REGION Network 339: CARRIER SPACING FAULT
   RUNG wire#powerrail
      Contact( "reset" )
      Contact( "EMS".Carrier[59].SDC_OUT.Faults.CarrierSpacingFault )
      wire#w1
      Coil( "DB302_HMI_Faults".Carrier59_Faults_2.%X2 )
   END_RUNG
   RUNG wire#powerrail
      Contact( "DB302_HMI_Faults".Carrier59_Faults_2.%X2 )
      I_Contact( "EMS_Fault_Reset" )
   END_RUNG wire#w1
   // the same network as SCL:
   "DB302_HMI_Faults".Carrier59_Faults_2.%X2 := ("reset" AND "EMS".Carrier[59].SDC_OUT.Faults.CarrierSpacingFault) OR ("DB302_HMI_Faults".Carrier59_Faults_2.%X2 AND NOT "EMS_Fault_Reset");
END_REGION

REGION Network 340: DUPLICATE CARRIER NUMBER FAULT
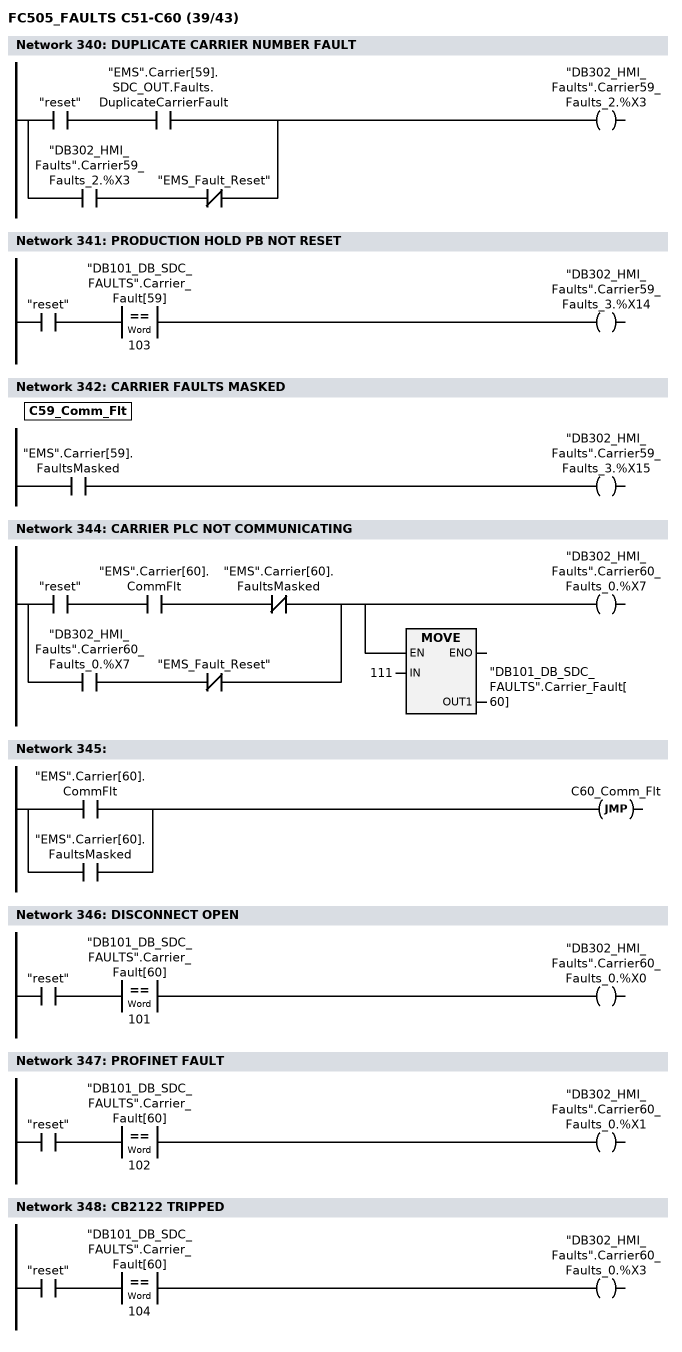
   RUNG wire#powerrail
      Contact( "reset" )
      Contact( "EMS".Carrier[59].SDC_OUT.Faults.DuplicateCarrierFault )
      wire#w1
      Coil( "DB302_HMI_Faults".Carrier59_Faults_2.%X3 )
   END_RUNG
   RUNG wire#powerrail
      Contact( "DB302_HMI_Faults".Carrier59_Faults_2.%X3 )
      I_Contact( "EMS_Fault_Reset" )
   END_RUNG wire#w1
   // the same network as SCL:
   "DB302_HMI_Faults".Carrier59_Faults_2.%X3 := ("reset" AND "EMS".Carrier[59].SDC_OUT.Faults.DuplicateCarrierFault) OR ("DB302_HMI_Faults".Carrier59_Faults_2.%X3 AND NOT "EMS_Fault_Reset");
END_REGION

REGION Network 341: PRODUCTION HOLD PB NOT RESET
   RUNG wire#powerrail
      Contact( "reset" )
      { S7_Templates := "SrcType := Word" } EQ_Contact(in1 := "DB101_DB_SDC_FAULTS".Carrier_Fault[59], in2 := 103)
      Coil( "DB302_HMI_Faults".Carrier59_Faults_3.%X14 )
   END_RUNG
   // the same network as SCL:
   "DB302_HMI_Faults".Carrier59_Faults_3.%X14 := "reset" AND ("DB101_DB_SDC_FAULTS".Carrier_Fault[59] = 103);
END_REGION

REGION Network 342: CARRIER FAULTS MASKED
   Label( C59_Comm_Flt )
   RUNG wire#powerrail
      Contact( "EMS".Carrier[59].FaultsMasked )
      Coil( "DB302_HMI_Faults".Carrier59_Faults_3.%X15 )
   END_RUNG
   // the same network as SCL:
   C59_Comm_Flt:
   "DB302_HMI_Faults".Carrier59_Faults_3.%X15 := "EMS".Carrier[59].FaultsMasked;
END_REGION

REGION Network 343: CARRIER 60 FAULTS
END_REGION

REGION Network 344: CARRIER PLC NOT COMMUNICATING
   RUNG wire#powerrail
      Contact( "reset" )
      Contact( "EMS".Carrier[60].CommFlt )
      I_Contact( "EMS".Carrier[60].FaultsMasked )
      wire#w1
      Coil( "DB302_HMI_Faults".Carrier60_Faults_0.%X7 )
   END_RUNG
   RUNG wire#powerrail
      Contact( "DB302_HMI_Faults".Carrier60_Faults_0.%X7 )
      I_Contact( "EMS_Fault_Reset" )
   END_RUNG wire#w1
   RUNG wire#w1
      Move(in := 111, out1 => "DB101_DB_SDC_FAULTS".Carrier_Fault[60])
   END_RUNG
   // the same network as SCL:
   "DB302_HMI_Faults".Carrier60_Faults_0.%X7 := ("reset" AND "EMS".Carrier[60].CommFlt AND NOT "EMS".Carrier[60].FaultsMasked) OR ("DB302_HMI_Faults".Carrier60_Faults_0.%X7 AND NOT "EMS_Fault_Reset");
   IF "DB302_HMI_Faults".Carrier60_Faults_0.%X7 THEN "DB101_DB_SDC_FAULTS".Carrier_Fault[60] := 111; END_IF;
END_REGION

REGION Network 345
   RUNG wire#powerrail
      Contact( "EMS".Carrier[60].CommFlt )
      wire#w1
      JumpCoil( C60_Comm_Flt )
   END_RUNG
   RUNG wire#powerrail
      Contact( "EMS".Carrier[60].FaultsMasked )
   END_RUNG wire#w1
   // the same network as SCL:
   IF "EMS".Carrier[60].CommFlt OR "EMS".Carrier[60].FaultsMasked THEN GOTO C60_Comm_Flt; END_IF;
END_REGION

REGION Network 346: DISCONNECT OPEN
   RUNG wire#powerrail
      Contact( "reset" )
      { S7_Templates := "SrcType := Word" } EQ_Contact(in1 := "DB101_DB_SDC_FAULTS".Carrier_Fault[60], in2 := 101)
      Coil( "DB302_HMI_Faults".Carrier60_Faults_0.%X0 )
   END_RUNG
   // the same network as SCL:
   "DB302_HMI_Faults".Carrier60_Faults_0.%X0 := "reset" AND ("DB101_DB_SDC_FAULTS".Carrier_Fault[60] = 101);
END_REGION

REGION Network 347: PROFINET FAULT
   RUNG wire#powerrail
      Contact( "reset" )
      { S7_Templates := "SrcType := Word" } EQ_Contact(in1 := "DB101_DB_SDC_FAULTS".Carrier_Fault[60], in2 := 102)
      Coil( "DB302_HMI_Faults".Carrier60_Faults_0.%X1 )
   END_RUNG
   // the same network as SCL:
   "DB302_HMI_Faults".Carrier60_Faults_0.%X1 := "reset" AND ("DB101_DB_SDC_FAULTS".Carrier_Fault[60] = 102);
END_REGION

REGION Network 348: CB2122 TRIPPED
   RUNG wire#powerrail
      Contact( "reset" )
      { S7_Templates := "SrcType := Word" } EQ_Contact(in1 := "DB101_DB_SDC_FAULTS".Carrier_Fault[60], in2 := 104)
      Coil( "DB302_HMI_Faults".Carrier60_Faults_0.%X3 )
   END_RUNG
   // the same network as SCL:
   "DB302_HMI_Faults".Carrier60_Faults_0.%X3 := "reset" AND ("DB101_DB_SDC_FAULTS".Carrier_Fault[60] = 104);
END_REGION

REGION Network 349: CB2123 TRIPPED
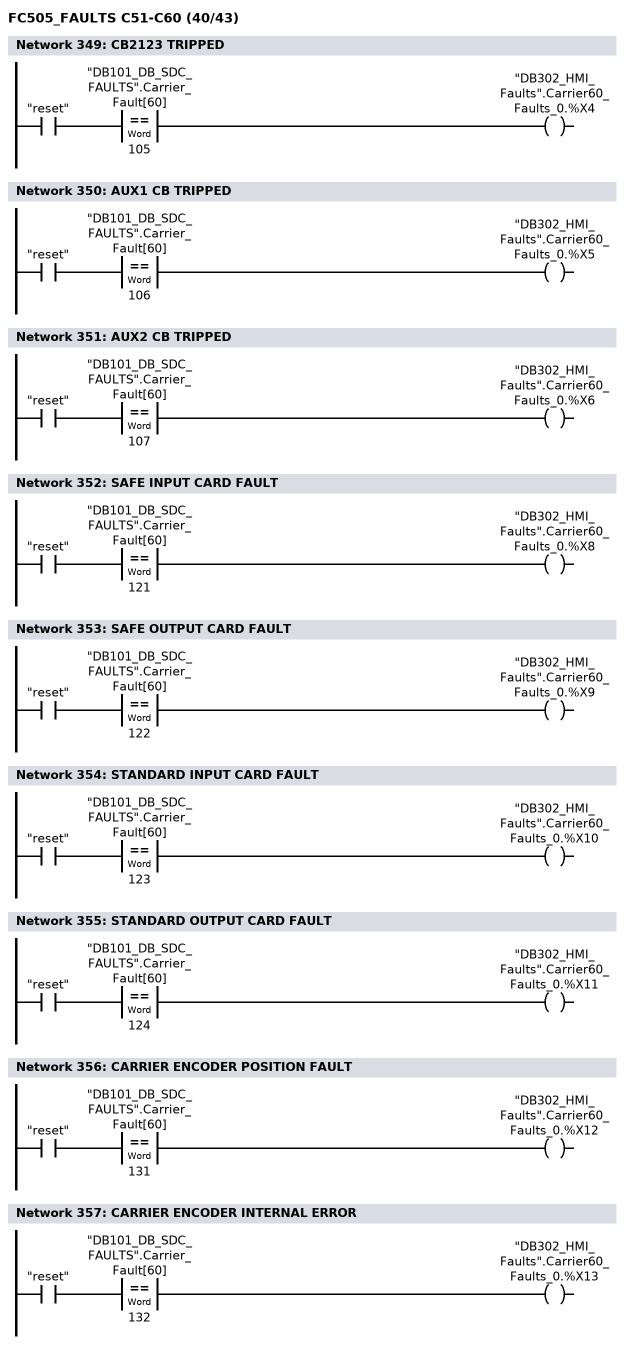
   RUNG wire#powerrail
      Contact( "reset" )
      { S7_Templates := "SrcType := Word" } EQ_Contact(in1 := "DB101_DB_SDC_FAULTS".Carrier_Fault[60], in2 := 105)
      Coil( "DB302_HMI_Faults".Carrier60_Faults_0.%X4 )
   END_RUNG
   // the same network as SCL:
   "DB302_HMI_Faults".Carrier60_Faults_0.%X4 := "reset" AND ("DB101_DB_SDC_FAULTS".Carrier_Fault[60] = 105);
END_REGION

REGION Network 350: AUX1 CB TRIPPED
   RUNG wire#powerrail
      Contact( "reset" )
      { S7_Templates := "SrcType := Word" } EQ_Contact(in1 := "DB101_DB_SDC_FAULTS".Carrier_Fault[60], in2 := 106)
      Coil( "DB302_HMI_Faults".Carrier60_Faults_0.%X5 )
   END_RUNG
   // the same network as SCL:
   "DB302_HMI_Faults".Carrier60_Faults_0.%X5 := "reset" AND ("DB101_DB_SDC_FAULTS".Carrier_Fault[60] = 106);
END_REGION

REGION Network 351: AUX2 CB TRIPPED
   RUNG wire#powerrail
      Contact( "reset" )
      { S7_Templates := "SrcType := Word" } EQ_Contact(in1 := "DB101_DB_SDC_FAULTS".Carrier_Fault[60], in2 := 107)
      Coil( "DB302_HMI_Faults".Carrier60_Faults_0.%X6 )
   END_RUNG
   // the same network as SCL:
   "DB302_HMI_Faults".Carrier60_Faults_0.%X6 := "reset" AND ("DB101_DB_SDC_FAULTS".Carrier_Fault[60] = 107);
END_REGION

REGION Network 352: SAFE INPUT CARD FAULT
   RUNG wire#powerrail
      Contact( "reset" )
      { S7_Templates := "SrcType := Word" } EQ_Contact(in1 := "DB101_DB_SDC_FAULTS".Carrier_Fault[60], in2 := 121)
      Coil( "DB302_HMI_Faults".Carrier60_Faults_0.%X8 )
   END_RUNG
   // the same network as SCL:
   "DB302_HMI_Faults".Carrier60_Faults_0.%X8 := "reset" AND ("DB101_DB_SDC_FAULTS".Carrier_Fault[60] = 121);
END_REGION

REGION Network 353: SAFE OUTPUT CARD FAULT
   RUNG wire#powerrail
      Contact( "reset" )
      { S7_Templates := "SrcType := Word" } EQ_Contact(in1 := "DB101_DB_SDC_FAULTS".Carrier_Fault[60], in2 := 122)
      Coil( "DB302_HMI_Faults".Carrier60_Faults_0.%X9 )
   END_RUNG
   // the same network as SCL:
   "DB302_HMI_Faults".Carrier60_Faults_0.%X9 := "reset" AND ("DB101_DB_SDC_FAULTS".Carrier_Fault[60] = 122);
END_REGION

REGION Network 354: STANDARD INPUT CARD FAULT
   RUNG wire#powerrail
      Contact( "reset" )
      { S7_Templates := "SrcType := Word" } EQ_Contact(in1 := "DB101_DB_SDC_FAULTS".Carrier_Fault[60], in2 := 123)
      Coil( "DB302_HMI_Faults".Carrier60_Faults_0.%X10 )
   END_RUNG
   // the same network as SCL:
   "DB302_HMI_Faults".Carrier60_Faults_0.%X10 := "reset" AND ("DB101_DB_SDC_FAULTS".Carrier_Fault[60] = 123);
END_REGION

REGION Network 355: STANDARD OUTPUT CARD FAULT
   RUNG wire#powerrail
      Contact( "reset" )
      { S7_Templates := "SrcType := Word" } EQ_Contact(in1 := "DB101_DB_SDC_FAULTS".Carrier_Fault[60], in2 := 124)
      Coil( "DB302_HMI_Faults".Carrier60_Faults_0.%X11 )
   END_RUNG
   // the same network as SCL:
   "DB302_HMI_Faults".Carrier60_Faults_0.%X11 := "reset" AND ("DB101_DB_SDC_FAULTS".Carrier_Fault[60] = 124);
END_REGION

REGION Network 356: CARRIER ENCODER POSITION FAULT
   RUNG wire#powerrail
      Contact( "reset" )
      { S7_Templates := "SrcType := Word" } EQ_Contact(in1 := "DB101_DB_SDC_FAULTS".Carrier_Fault[60], in2 := 131)
      Coil( "DB302_HMI_Faults".Carrier60_Faults_0.%X12 )
   END_RUNG
   // the same network as SCL:
   "DB302_HMI_Faults".Carrier60_Faults_0.%X12 := "reset" AND ("DB101_DB_SDC_FAULTS".Carrier_Fault[60] = 131);
END_REGION

REGION Network 357: CARRIER ENCODER INTERNAL ERROR
   RUNG wire#powerrail
      Contact( "reset" )
      { S7_Templates := "SrcType := Word" } EQ_Contact(in1 := "DB101_DB_SDC_FAULTS".Carrier_Fault[60], in2 := 132)
      Coil( "DB302_HMI_Faults".Carrier60_Faults_0.%X13 )
   END_RUNG
   // the same network as SCL:
   "DB302_HMI_Faults".Carrier60_Faults_0.%X13 := "reset" AND ("DB101_DB_SDC_FAULTS".Carrier_Fault[60] = 132);
END_REGION

REGION Network 358: CARRIER ENCODER COMM FAULT
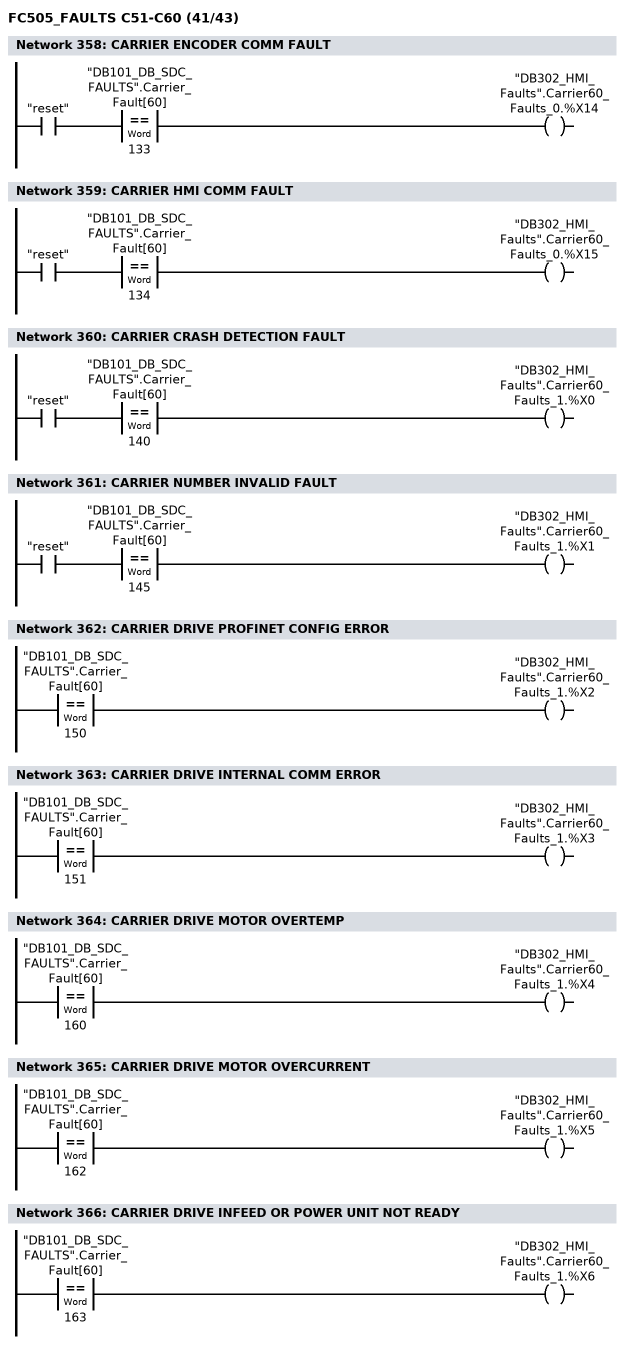
   RUNG wire#powerrail
      Contact( "reset" )
      { S7_Templates := "SrcType := Word" } EQ_Contact(in1 := "DB101_DB_SDC_FAULTS".Carrier_Fault[60], in2 := 133)
      Coil( "DB302_HMI_Faults".Carrier60_Faults_0.%X14 )
   END_RUNG
   // the same network as SCL:
   "DB302_HMI_Faults".Carrier60_Faults_0.%X14 := "reset" AND ("DB101_DB_SDC_FAULTS".Carrier_Fault[60] = 133);
END_REGION

REGION Network 359: CARRIER HMI COMM FAULT
   RUNG wire#powerrail
      Contact( "reset" )
      { S7_Templates := "SrcType := Word" } EQ_Contact(in1 := "DB101_DB_SDC_FAULTS".Carrier_Fault[60], in2 := 134)
      Coil( "DB302_HMI_Faults".Carrier60_Faults_0.%X15 )
   END_RUNG
   // the same network as SCL:
   "DB302_HMI_Faults".Carrier60_Faults_0.%X15 := "reset" AND ("DB101_DB_SDC_FAULTS".Carrier_Fault[60] = 134);
END_REGION

REGION Network 360: CARRIER CRASH DETECTION FAULT
   RUNG wire#powerrail
      Contact( "reset" )
      { S7_Templates := "SrcType := Word" } EQ_Contact(in1 := "DB101_DB_SDC_FAULTS".Carrier_Fault[60], in2 := 140)
      Coil( "DB302_HMI_Faults".Carrier60_Faults_1.%X0 )
   END_RUNG
   // the same network as SCL:
   "DB302_HMI_Faults".Carrier60_Faults_1.%X0 := "reset" AND ("DB101_DB_SDC_FAULTS".Carrier_Fault[60] = 140);
END_REGION

REGION Network 361: CARRIER NUMBER INVALID FAULT
   RUNG wire#powerrail
      Contact( "reset" )
      { S7_Templates := "SrcType := Word" } EQ_Contact(in1 := "DB101_DB_SDC_FAULTS".Carrier_Fault[60], in2 := 145)
      Coil( "DB302_HMI_Faults".Carrier60_Faults_1.%X1 )
   END_RUNG
   // the same network as SCL:
   "DB302_HMI_Faults".Carrier60_Faults_1.%X1 := "reset" AND ("DB101_DB_SDC_FAULTS".Carrier_Fault[60] = 145);
END_REGION

REGION Network 362: CARRIER DRIVE PROFINET CONFIG ERROR
   RUNG wire#powerrail
      { S7_Templates := "SrcType := Word" } EQ_Contact(in1 := "DB101_DB_SDC_FAULTS".Carrier_Fault[60], in2 := 150)
      Coil( "DB302_HMI_Faults".Carrier60_Faults_1.%X2 )
   END_RUNG
   // the same network as SCL:
   "DB302_HMI_Faults".Carrier60_Faults_1.%X2 := "DB101_DB_SDC_FAULTS".Carrier_Fault[60] = 150;
END_REGION

REGION Network 363: CARRIER DRIVE INTERNAL COMM ERROR
   RUNG wire#powerrail
      { S7_Templates := "SrcType := Word" } EQ_Contact(in1 := "DB101_DB_SDC_FAULTS".Carrier_Fault[60], in2 := 151)
      Coil( "DB302_HMI_Faults".Carrier60_Faults_1.%X3 )
   END_RUNG
   // the same network as SCL:
   "DB302_HMI_Faults".Carrier60_Faults_1.%X3 := "DB101_DB_SDC_FAULTS".Carrier_Fault[60] = 151;
END_REGION

REGION Network 364: CARRIER DRIVE MOTOR OVERTEMP
   RUNG wire#powerrail
      { S7_Templates := "SrcType := Word" } EQ_Contact(in1 := "DB101_DB_SDC_FAULTS".Carrier_Fault[60], in2 := 160)
      Coil( "DB302_HMI_Faults".Carrier60_Faults_1.%X4 )
   END_RUNG
   // the same network as SCL:
   "DB302_HMI_Faults".Carrier60_Faults_1.%X4 := "DB101_DB_SDC_FAULTS".Carrier_Fault[60] = 160;
END_REGION

REGION Network 365: CARRIER DRIVE MOTOR OVERCURRENT
   RUNG wire#powerrail
      { S7_Templates := "SrcType := Word" } EQ_Contact(in1 := "DB101_DB_SDC_FAULTS".Carrier_Fault[60], in2 := 162)
      Coil( "DB302_HMI_Faults".Carrier60_Faults_1.%X5 )
   END_RUNG
   // the same network as SCL:
   "DB302_HMI_Faults".Carrier60_Faults_1.%X5 := "DB101_DB_SDC_FAULTS".Carrier_Fault[60] = 162;
END_REGION

REGION Network 366: CARRIER DRIVE INFEED OR POWER UNIT NOT READY
   RUNG wire#powerrail
      { S7_Templates := "SrcType := Word" } EQ_Contact(in1 := "DB101_DB_SDC_FAULTS".Carrier_Fault[60], in2 := 163)
      Coil( "DB302_HMI_Faults".Carrier60_Faults_1.%X6 )
   END_RUNG
   // the same network as SCL:
   "DB302_HMI_Faults".Carrier60_Faults_1.%X6 := "DB101_DB_SDC_FAULTS".Carrier_Fault[60] = 163;
END_REGION

REGION Network 367: CARRIER DRIVE SHORT CIRCUIT / GROUND FAULT DETECTED
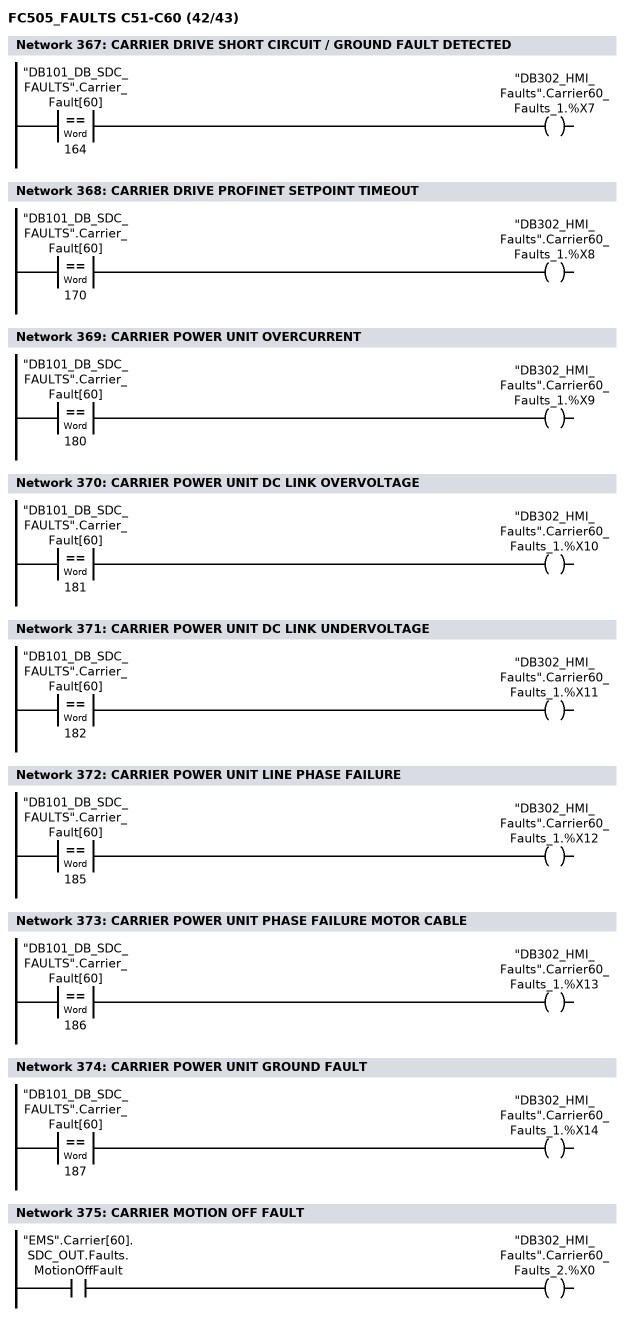
   RUNG wire#powerrail
      { S7_Templates := "SrcType := Word" } EQ_Contact(in1 := "DB101_DB_SDC_FAULTS".Carrier_Fault[60], in2 := 164)
      Coil( "DB302_HMI_Faults".Carrier60_Faults_1.%X7 )
   END_RUNG
   // the same network as SCL:
   "DB302_HMI_Faults".Carrier60_Faults_1.%X7 := "DB101_DB_SDC_FAULTS".Carrier_Fault[60] = 164;
END_REGION

REGION Network 368: CARRIER DRIVE PROFINET SETPOINT TIMEOUT
   RUNG wire#powerrail
      { S7_Templates := "SrcType := Word" } EQ_Contact(in1 := "DB101_DB_SDC_FAULTS".Carrier_Fault[60], in2 := 170)
      Coil( "DB302_HMI_Faults".Carrier60_Faults_1.%X8 )
   END_RUNG
   // the same network as SCL:
   "DB302_HMI_Faults".Carrier60_Faults_1.%X8 := "DB101_DB_SDC_FAULTS".Carrier_Fault[60] = 170;
END_REGION

REGION Network 369: CARRIER POWER UNIT OVERCURRENT
   RUNG wire#powerrail
      { S7_Templates := "SrcType := Word" } EQ_Contact(in1 := "DB101_DB_SDC_FAULTS".Carrier_Fault[60], in2 := 180)
      Coil( "DB302_HMI_Faults".Carrier60_Faults_1.%X9 )
   END_RUNG
   // the same network as SCL:
   "DB302_HMI_Faults".Carrier60_Faults_1.%X9 := "DB101_DB_SDC_FAULTS".Carrier_Fault[60] = 180;
END_REGION

REGION Network 370: CARRIER POWER UNIT DC LINK OVERVOLTAGE
   RUNG wire#powerrail
      { S7_Templates := "SrcType := Word" } EQ_Contact(in1 := "DB101_DB_SDC_FAULTS".Carrier_Fault[60], in2 := 181)
      Coil( "DB302_HMI_Faults".Carrier60_Faults_1.%X10 )
   END_RUNG
   // the same network as SCL:
   "DB302_HMI_Faults".Carrier60_Faults_1.%X10 := "DB101_DB_SDC_FAULTS".Carrier_Fault[60] = 181;
END_REGION

REGION Network 371: CARRIER POWER UNIT DC LINK UNDERVOLTAGE
   RUNG wire#powerrail
      { S7_Templates := "SrcType := Word" } EQ_Contact(in1 := "DB101_DB_SDC_FAULTS".Carrier_Fault[60], in2 := 182)
      Coil( "DB302_HMI_Faults".Carrier60_Faults_1.%X11 )
   END_RUNG
   // the same network as SCL:
   "DB302_HMI_Faults".Carrier60_Faults_1.%X11 := "DB101_DB_SDC_FAULTS".Carrier_Fault[60] = 182;
END_REGION

REGION Network 372: CARRIER POWER UNIT LINE PHASE FAILURE
   RUNG wire#powerrail
      { S7_Templates := "SrcType := Word" } EQ_Contact(in1 := "DB101_DB_SDC_FAULTS".Carrier_Fault[60], in2 := 185)
      Coil( "DB302_HMI_Faults".Carrier60_Faults_1.%X12 )
   END_RUNG
   // the same network as SCL:
   "DB302_HMI_Faults".Carrier60_Faults_1.%X12 := "DB101_DB_SDC_FAULTS".Carrier_Fault[60] = 185;
END_REGION

REGION Network 373: CARRIER POWER UNIT PHASE FAILURE MOTOR CABLE
   RUNG wire#powerrail
      { S7_Templates := "SrcType := Word" } EQ_Contact(in1 := "DB101_DB_SDC_FAULTS".Carrier_Fault[60], in2 := 186)
      Coil( "DB302_HMI_Faults".Carrier60_Faults_1.%X13 )
   END_RUNG
   // the same network as SCL:
   "DB302_HMI_Faults".Carrier60_Faults_1.%X13 := "DB101_DB_SDC_FAULTS".Carrier_Fault[60] = 186;
END_REGION

REGION Network 374: CARRIER POWER UNIT GROUND FAULT
   RUNG wire#powerrail
      { S7_Templates := "SrcType := Word" } EQ_Contact(in1 := "DB101_DB_SDC_FAULTS".Carrier_Fault[60], in2 := 187)
      Coil( "DB302_HMI_Faults".Carrier60_Faults_1.%X14 )
   END_RUNG
   // the same network as SCL:
   "DB302_HMI_Faults".Carrier60_Faults_1.%X14 := "DB101_DB_SDC_FAULTS".Carrier_Fault[60] = 187;
END_REGION

REGION Network 375: CARRIER MOTION OFF FAULT
   RUNG wire#powerrail
      Contact( "EMS".Carrier[60].SDC_OUT.Faults.MotionOffFault )
      Coil( "DB302_HMI_Faults".Carrier60_Faults_2.%X0 )
   END_RUNG
   // the same network as SCL:
   "DB302_HMI_Faults".Carrier60_Faults_2.%X0 := "EMS".Carrier[60].SDC_OUT.Faults.MotionOffFault;
END_REGION

REGION Network 376: CARRIER MOTION ON FAULT
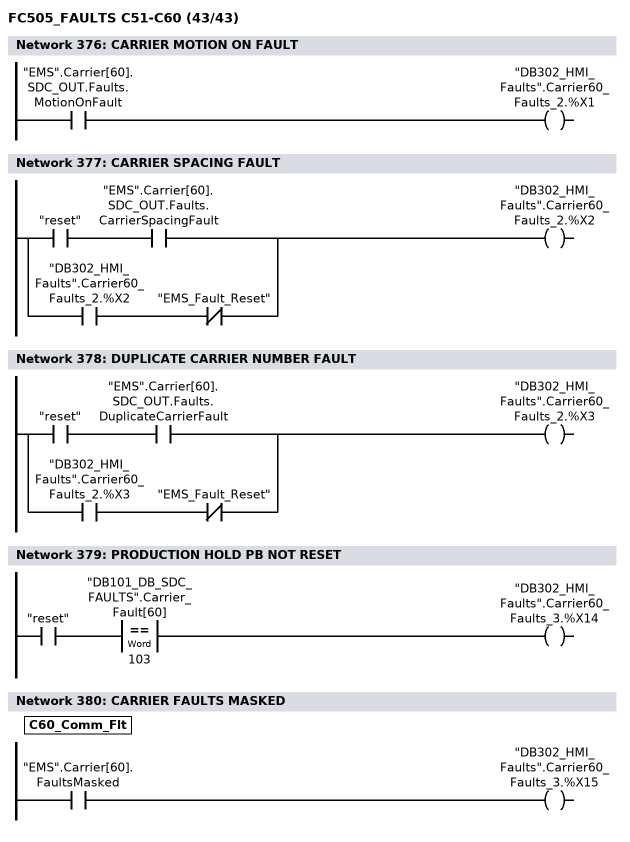
   RUNG wire#powerrail
      Contact( "EMS".Carrier[60].SDC_OUT.Faults.MotionOnFault )
      Coil( "DB302_HMI_Faults".Carrier60_Faults_2.%X1 )
   END_RUNG
   // the same network as SCL:
   "DB302_HMI_Faults".Carrier60_Faults_2.%X1 := "EMS".Carrier[60].SDC_OUT.Faults.MotionOnFault;
END_REGION

REGION Network 377: CARRIER SPACING FAULT
   RUNG wire#powerrail
      Contact( "reset" )
      Contact( "EMS".Carrier[60].SDC_OUT.Faults.CarrierSpacingFault )
      wire#w1
      Coil( "DB302_HMI_Faults".Carrier60_Faults_2.%X2 )
   END_RUNG
   RUNG wire#powerrail
      Contact( "DB302_HMI_Faults".Carrier60_Faults_2.%X2 )
      I_Contact( "EMS_Fault_Reset" )
   END_RUNG wire#w1
   // the same network as SCL:
   "DB302_HMI_Faults".Carrier60_Faults_2.%X2 := ("reset" AND "EMS".Carrier[60].SDC_OUT.Faults.CarrierSpacingFault) OR ("DB302_HMI_Faults".Carrier60_Faults_2.%X2 AND NOT "EMS_Fault_Reset");
END_REGION

REGION Network 378: DUPLICATE CARRIER NUMBER FAULT
   RUNG wire#powerrail
      Contact( "reset" )
      Contact( "EMS".Carrier[60].SDC_OUT.Faults.DuplicateCarrierFault )
      wire#w1
      Coil( "DB302_HMI_Faults".Carrier60_Faults_2.%X3 )
   END_RUNG
   RUNG wire#powerrail
      Contact( "DB302_HMI_Faults".Carrier60_Faults_2.%X3 )
      I_Contact( "EMS_Fault_Reset" )
   END_RUNG wire#w1
   // the same network as SCL:
   "DB302_HMI_Faults".Carrier60_Faults_2.%X3 := ("reset" AND "EMS".Carrier[60].SDC_OUT.Faults.DuplicateCarrierFault) OR ("DB302_HMI_Faults".Carrier60_Faults_2.%X3 AND NOT "EMS_Fault_Reset");
END_REGION

REGION Network 379: PRODUCTION HOLD PB NOT RESET
   RUNG wire#powerrail
      Contact( "reset" )
      { S7_Templates := "SrcType := Word" } EQ_Contact(in1 := "DB101_DB_SDC_FAULTS".Carrier_Fault[60], in2 := 103)
      Coil( "DB302_HMI_Faults".Carrier60_Faults_3.%X14 )
   END_RUNG
   // the same network as SCL:
   "DB302_HMI_Faults".Carrier60_Faults_3.%X14 := "reset" AND ("DB101_DB_SDC_FAULTS".Carrier_Fault[60] = 103);
END_REGION

REGION Network 380: CARRIER FAULTS MASKED
   Label( C60_Comm_Flt )
   RUNG wire#powerrail
      Contact( "EMS".Carrier[60].FaultsMasked )
      Coil( "DB302_HMI_Faults".Carrier60_Faults_3.%X15 )
   END_RUNG
   // the same network as SCL:
   C60_Comm_Flt:
   "DB302_HMI_Faults".Carrier60_Faults_3.%X15 := "EMS".Carrier[60].FaultsMasked;
END_REGION
END_FUNCTION

FUNCTION "FC506_FAULTS C61-C70" : Void   // FC506, LAD
{ S7_Optimized_Access := 'TRUE' }
VERSION : 0.1
BEGIN

REGION Network 1: CARRIER 61 FAULTS
END_REGION

REGION Network 2: CARRIER PLC NOT COMMUNICATING
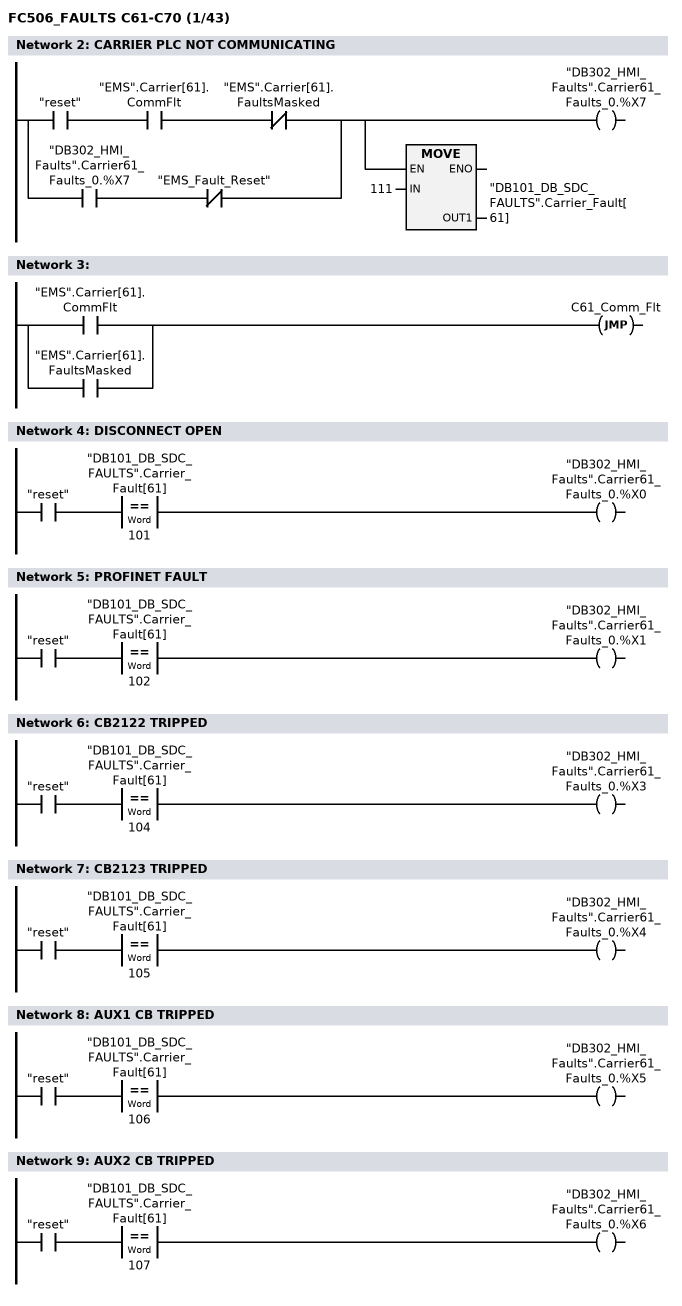
   RUNG wire#powerrail
      Contact( "reset" )
      Contact( "EMS".Carrier[61].CommFlt )
      I_Contact( "EMS".Carrier[61].FaultsMasked )
      wire#w1
      Coil( "DB302_HMI_Faults".Carrier61_Faults_0.%X7 )
   END_RUNG
   RUNG wire#powerrail
      Contact( "DB302_HMI_Faults".Carrier61_Faults_0.%X7 )
      I_Contact( "EMS_Fault_Reset" )
   END_RUNG wire#w1
   RUNG wire#w1
      Move(in := 111, out1 => "DB101_DB_SDC_FAULTS".Carrier_Fault[61])
   END_RUNG
   // the same network as SCL:
   "DB302_HMI_Faults".Carrier61_Faults_0.%X7 := ("reset" AND "EMS".Carrier[61].CommFlt AND NOT "EMS".Carrier[61].FaultsMasked) OR ("DB302_HMI_Faults".Carrier61_Faults_0.%X7 AND NOT "EMS_Fault_Reset");
   IF "DB302_HMI_Faults".Carrier61_Faults_0.%X7 THEN "DB101_DB_SDC_FAULTS".Carrier_Fault[61] := 111; END_IF;
END_REGION

REGION Network 3
   RUNG wire#powerrail
      Contact( "EMS".Carrier[61].CommFlt )
      wire#w1
      JumpCoil( C61_Comm_Flt )
   END_RUNG
   RUNG wire#powerrail
      Contact( "EMS".Carrier[61].FaultsMasked )
   END_RUNG wire#w1
   // the same network as SCL:
   IF "EMS".Carrier[61].CommFlt OR "EMS".Carrier[61].FaultsMasked THEN GOTO C61_Comm_Flt; END_IF;
END_REGION

REGION Network 4: DISCONNECT OPEN
   RUNG wire#powerrail
      Contact( "reset" )
      { S7_Templates := "SrcType := Word" } EQ_Contact(in1 := "DB101_DB_SDC_FAULTS".Carrier_Fault[61], in2 := 101)
      Coil( "DB302_HMI_Faults".Carrier61_Faults_0.%X0 )
   END_RUNG
   // the same network as SCL:
   "DB302_HMI_Faults".Carrier61_Faults_0.%X0 := "reset" AND ("DB101_DB_SDC_FAULTS".Carrier_Fault[61] = 101);
END_REGION

REGION Network 5: PROFINET FAULT
   RUNG wire#powerrail
      Contact( "reset" )
      { S7_Templates := "SrcType := Word" } EQ_Contact(in1 := "DB101_DB_SDC_FAULTS".Carrier_Fault[61], in2 := 102)
      Coil( "DB302_HMI_Faults".Carrier61_Faults_0.%X1 )
   END_RUNG
   // the same network as SCL:
   "DB302_HMI_Faults".Carrier61_Faults_0.%X1 := "reset" AND ("DB101_DB_SDC_FAULTS".Carrier_Fault[61] = 102);
END_REGION

REGION Network 6: CB2122 TRIPPED
   RUNG wire#powerrail
      Contact( "reset" )
      { S7_Templates := "SrcType := Word" } EQ_Contact(in1 := "DB101_DB_SDC_FAULTS".Carrier_Fault[61], in2 := 104)
      Coil( "DB302_HMI_Faults".Carrier61_Faults_0.%X3 )
   END_RUNG
   // the same network as SCL:
   "DB302_HMI_Faults".Carrier61_Faults_0.%X3 := "reset" AND ("DB101_DB_SDC_FAULTS".Carrier_Fault[61] = 104);
END_REGION

REGION Network 7: CB2123 TRIPPED
   RUNG wire#powerrail
      Contact( "reset" )
      { S7_Templates := "SrcType := Word" } EQ_Contact(in1 := "DB101_DB_SDC_FAULTS".Carrier_Fault[61], in2 := 105)
      Coil( "DB302_HMI_Faults".Carrier61_Faults_0.%X4 )
   END_RUNG
   // the same network as SCL:
   "DB302_HMI_Faults".Carrier61_Faults_0.%X4 := "reset" AND ("DB101_DB_SDC_FAULTS".Carrier_Fault[61] = 105);
END_REGION

REGION Network 8: AUX1 CB TRIPPED
   RUNG wire#powerrail
      Contact( "reset" )
      { S7_Templates := "SrcType := Word" } EQ_Contact(in1 := "DB101_DB_SDC_FAULTS".Carrier_Fault[61], in2 := 106)
      Coil( "DB302_HMI_Faults".Carrier61_Faults_0.%X5 )
   END_RUNG
   // the same network as SCL:
   "DB302_HMI_Faults".Carrier61_Faults_0.%X5 := "reset" AND ("DB101_DB_SDC_FAULTS".Carrier_Fault[61] = 106);
END_REGION

REGION Network 9: AUX2 CB TRIPPED
   RUNG wire#powerrail
      Contact( "reset" )
      { S7_Templates := "SrcType := Word" } EQ_Contact(in1 := "DB101_DB_SDC_FAULTS".Carrier_Fault[61], in2 := 107)
      Coil( "DB302_HMI_Faults".Carrier61_Faults_0.%X6 )
   END_RUNG
   // the same network as SCL:
   "DB302_HMI_Faults".Carrier61_Faults_0.%X6 := "reset" AND ("DB101_DB_SDC_FAULTS".Carrier_Fault[61] = 107);
END_REGION

REGION Network 10: SAFE INPUT CARD FAULT
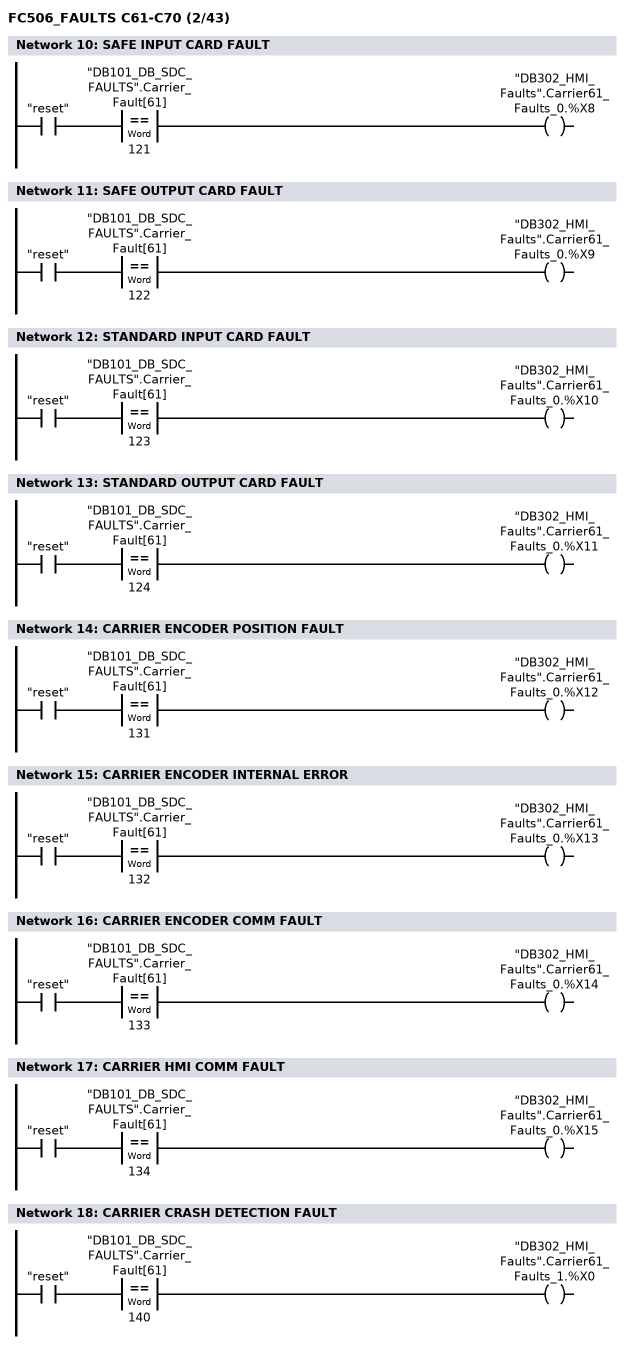
   RUNG wire#powerrail
      Contact( "reset" )
      { S7_Templates := "SrcType := Word" } EQ_Contact(in1 := "DB101_DB_SDC_FAULTS".Carrier_Fault[61], in2 := 121)
      Coil( "DB302_HMI_Faults".Carrier61_Faults_0.%X8 )
   END_RUNG
   // the same network as SCL:
   "DB302_HMI_Faults".Carrier61_Faults_0.%X8 := "reset" AND ("DB101_DB_SDC_FAULTS".Carrier_Fault[61] = 121);
END_REGION

REGION Network 11: SAFE OUTPUT CARD FAULT
   RUNG wire#powerrail
      Contact( "reset" )
      { S7_Templates := "SrcType := Word" } EQ_Contact(in1 := "DB101_DB_SDC_FAULTS".Carrier_Fault[61], in2 := 122)
      Coil( "DB302_HMI_Faults".Carrier61_Faults_0.%X9 )
   END_RUNG
   // the same network as SCL:
   "DB302_HMI_Faults".Carrier61_Faults_0.%X9 := "reset" AND ("DB101_DB_SDC_FAULTS".Carrier_Fault[61] = 122);
END_REGION

REGION Network 12: STANDARD INPUT CARD FAULT
   RUNG wire#powerrail
      Contact( "reset" )
      { S7_Templates := "SrcType := Word" } EQ_Contact(in1 := "DB101_DB_SDC_FAULTS".Carrier_Fault[61], in2 := 123)
      Coil( "DB302_HMI_Faults".Carrier61_Faults_0.%X10 )
   END_RUNG
   // the same network as SCL:
   "DB302_HMI_Faults".Carrier61_Faults_0.%X10 := "reset" AND ("DB101_DB_SDC_FAULTS".Carrier_Fault[61] = 123);
END_REGION

REGION Network 13: STANDARD OUTPUT CARD FAULT
   RUNG wire#powerrail
      Contact( "reset" )
      { S7_Templates := "SrcType := Word" } EQ_Contact(in1 := "DB101_DB_SDC_FAULTS".Carrier_Fault[61], in2 := 124)
      Coil( "DB302_HMI_Faults".Carrier61_Faults_0.%X11 )
   END_RUNG
   // the same network as SCL:
   "DB302_HMI_Faults".Carrier61_Faults_0.%X11 := "reset" AND ("DB101_DB_SDC_FAULTS".Carrier_Fault[61] = 124);
END_REGION

REGION Network 14: CARRIER ENCODER POSITION FAULT
   RUNG wire#powerrail
      Contact( "reset" )
      { S7_Templates := "SrcType := Word" } EQ_Contact(in1 := "DB101_DB_SDC_FAULTS".Carrier_Fault[61], in2 := 131)
      Coil( "DB302_HMI_Faults".Carrier61_Faults_0.%X12 )
   END_RUNG
   // the same network as SCL:
   "DB302_HMI_Faults".Carrier61_Faults_0.%X12 := "reset" AND ("DB101_DB_SDC_FAULTS".Carrier_Fault[61] = 131);
END_REGION

REGION Network 15: CARRIER ENCODER INTERNAL ERROR
   RUNG wire#powerrail
      Contact( "reset" )
      { S7_Templates := "SrcType := Word" } EQ_Contact(in1 := "DB101_DB_SDC_FAULTS".Carrier_Fault[61], in2 := 132)
      Coil( "DB302_HMI_Faults".Carrier61_Faults_0.%X13 )
   END_RUNG
   // the same network as SCL:
   "DB302_HMI_Faults".Carrier61_Faults_0.%X13 := "reset" AND ("DB101_DB_SDC_FAULTS".Carrier_Fault[61] = 132);
END_REGION

REGION Network 16: CARRIER ENCODER COMM FAULT
   RUNG wire#powerrail
      Contact( "reset" )
      { S7_Templates := "SrcType := Word" } EQ_Contact(in1 := "DB101_DB_SDC_FAULTS".Carrier_Fault[61], in2 := 133)
      Coil( "DB302_HMI_Faults".Carrier61_Faults_0.%X14 )
   END_RUNG
   // the same network as SCL:
   "DB302_HMI_Faults".Carrier61_Faults_0.%X14 := "reset" AND ("DB101_DB_SDC_FAULTS".Carrier_Fault[61] = 133);
END_REGION

REGION Network 17: CARRIER HMI COMM FAULT
   RUNG wire#powerrail
      Contact( "reset" )
      { S7_Templates := "SrcType := Word" } EQ_Contact(in1 := "DB101_DB_SDC_FAULTS".Carrier_Fault[61], in2 := 134)
      Coil( "DB302_HMI_Faults".Carrier61_Faults_0.%X15 )
   END_RUNG
   // the same network as SCL:
   "DB302_HMI_Faults".Carrier61_Faults_0.%X15 := "reset" AND ("DB101_DB_SDC_FAULTS".Carrier_Fault[61] = 134);
END_REGION

REGION Network 18: CARRIER CRASH DETECTION FAULT
   RUNG wire#powerrail
      Contact( "reset" )
      { S7_Templates := "SrcType := Word" } EQ_Contact(in1 := "DB101_DB_SDC_FAULTS".Carrier_Fault[61], in2 := 140)
      Coil( "DB302_HMI_Faults".Carrier61_Faults_1.%X0 )
   END_RUNG
   // the same network as SCL:
   "DB302_HMI_Faults".Carrier61_Faults_1.%X0 := "reset" AND ("DB101_DB_SDC_FAULTS".Carrier_Fault[61] = 140);
END_REGION

REGION Network 19: CARRIER NUMBER INVALID FAULT
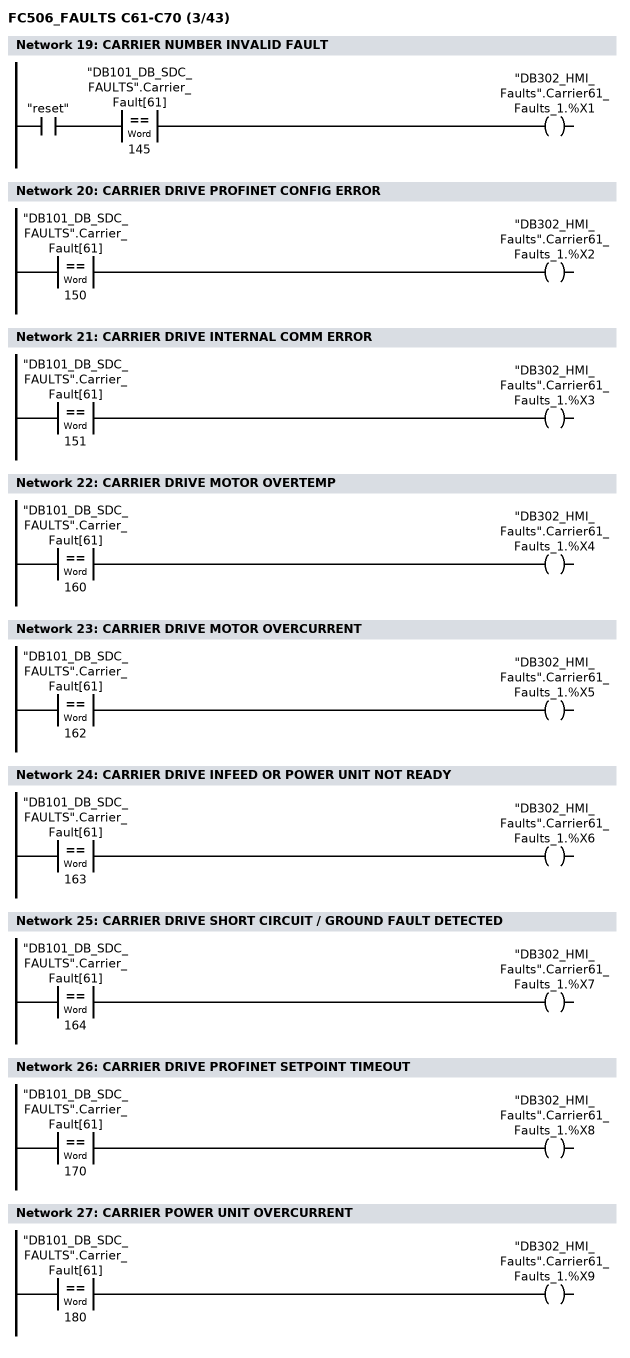
   RUNG wire#powerrail
      Contact( "reset" )
      { S7_Templates := "SrcType := Word" } EQ_Contact(in1 := "DB101_DB_SDC_FAULTS".Carrier_Fault[61], in2 := 145)
      Coil( "DB302_HMI_Faults".Carrier61_Faults_1.%X1 )
   END_RUNG
   // the same network as SCL:
   "DB302_HMI_Faults".Carrier61_Faults_1.%X1 := "reset" AND ("DB101_DB_SDC_FAULTS".Carrier_Fault[61] = 145);
END_REGION

REGION Network 20: CARRIER DRIVE PROFINET CONFIG ERROR
   RUNG wire#powerrail
      { S7_Templates := "SrcType := Word" } EQ_Contact(in1 := "DB101_DB_SDC_FAULTS".Carrier_Fault[61], in2 := 150)
      Coil( "DB302_HMI_Faults".Carrier61_Faults_1.%X2 )
   END_RUNG
   // the same network as SCL:
   "DB302_HMI_Faults".Carrier61_Faults_1.%X2 := "DB101_DB_SDC_FAULTS".Carrier_Fault[61] = 150;
END_REGION

REGION Network 21: CARRIER DRIVE INTERNAL COMM ERROR
   RUNG wire#powerrail
      { S7_Templates := "SrcType := Word" } EQ_Contact(in1 := "DB101_DB_SDC_FAULTS".Carrier_Fault[61], in2 := 151)
      Coil( "DB302_HMI_Faults".Carrier61_Faults_1.%X3 )
   END_RUNG
   // the same network as SCL:
   "DB302_HMI_Faults".Carrier61_Faults_1.%X3 := "DB101_DB_SDC_FAULTS".Carrier_Fault[61] = 151;
END_REGION

REGION Network 22: CARRIER DRIVE MOTOR OVERTEMP
   RUNG wire#powerrail
      { S7_Templates := "SrcType := Word" } EQ_Contact(in1 := "DB101_DB_SDC_FAULTS".Carrier_Fault[61], in2 := 160)
      Coil( "DB302_HMI_Faults".Carrier61_Faults_1.%X4 )
   END_RUNG
   // the same network as SCL:
   "DB302_HMI_Faults".Carrier61_Faults_1.%X4 := "DB101_DB_SDC_FAULTS".Carrier_Fault[61] = 160;
END_REGION

REGION Network 23: CARRIER DRIVE MOTOR OVERCURRENT
   RUNG wire#powerrail
      { S7_Templates := "SrcType := Word" } EQ_Contact(in1 := "DB101_DB_SDC_FAULTS".Carrier_Fault[61], in2 := 162)
      Coil( "DB302_HMI_Faults".Carrier61_Faults_1.%X5 )
   END_RUNG
   // the same network as SCL:
   "DB302_HMI_Faults".Carrier61_Faults_1.%X5 := "DB101_DB_SDC_FAULTS".Carrier_Fault[61] = 162;
END_REGION

REGION Network 24: CARRIER DRIVE INFEED OR POWER UNIT NOT READY
   RUNG wire#powerrail
      { S7_Templates := "SrcType := Word" } EQ_Contact(in1 := "DB101_DB_SDC_FAULTS".Carrier_Fault[61], in2 := 163)
      Coil( "DB302_HMI_Faults".Carrier61_Faults_1.%X6 )
   END_RUNG
   // the same network as SCL:
   "DB302_HMI_Faults".Carrier61_Faults_1.%X6 := "DB101_DB_SDC_FAULTS".Carrier_Fault[61] = 163;
END_REGION

REGION Network 25: CARRIER DRIVE SHORT CIRCUIT / GROUND FAULT DETECTED
   RUNG wire#powerrail
      { S7_Templates := "SrcType := Word" } EQ_Contact(in1 := "DB101_DB_SDC_FAULTS".Carrier_Fault[61], in2 := 164)
      Coil( "DB302_HMI_Faults".Carrier61_Faults_1.%X7 )
   END_RUNG
   // the same network as SCL:
   "DB302_HMI_Faults".Carrier61_Faults_1.%X7 := "DB101_DB_SDC_FAULTS".Carrier_Fault[61] = 164;
END_REGION

REGION Network 26: CARRIER DRIVE PROFINET SETPOINT TIMEOUT
   RUNG wire#powerrail
      { S7_Templates := "SrcType := Word" } EQ_Contact(in1 := "DB101_DB_SDC_FAULTS".Carrier_Fault[61], in2 := 170)
      Coil( "DB302_HMI_Faults".Carrier61_Faults_1.%X8 )
   END_RUNG
   // the same network as SCL:
   "DB302_HMI_Faults".Carrier61_Faults_1.%X8 := "DB101_DB_SDC_FAULTS".Carrier_Fault[61] = 170;
END_REGION

REGION Network 27: CARRIER POWER UNIT OVERCURRENT
   RUNG wire#powerrail
      { S7_Templates := "SrcType := Word" } EQ_Contact(in1 := "DB101_DB_SDC_FAULTS".Carrier_Fault[61], in2 := 180)
      Coil( "DB302_HMI_Faults".Carrier61_Faults_1.%X9 )
   END_RUNG
   // the same network as SCL:
   "DB302_HMI_Faults".Carrier61_Faults_1.%X9 := "DB101_DB_SDC_FAULTS".Carrier_Fault[61] = 180;
END_REGION

REGION Network 28: CARRIER POWER UNIT DC LINK OVERVOLTAGE